// TIA Portal project "maupTIA_DEMO2023_V17" (V17)

(* hardware
DEVICE "S71500/ET200MP station_1"  S7-1500 station
   slot 0: "Rail_0"  Rack  6ES7 590-1***0-0AA0
   slot 1: "PLC_1"  CPU 1512C-1 PN  6ES7 512-1CK00-0AB0  V2.1
      slot 3: "CPU display_1"  6ES7591-1AA00-0AA0
DEVICE "HMI_1"  TP700 Comfort
   slot 0: "TP700 Comfort"  TP700 Comfort  6AV2 124-0GC01-0AX0  14.0.1.0
   slot 1: "HMI_RT_1"  TP700 Comfort  6AV2 124-0GC01-0AX0  14.0.1.0
   slot 5: "HMI_1.IE_CP_1"  PROFINET Interface  14.0.1.0
      slot 1: "PROFINET Interface_1"  PROFINET Interface
         slot 1: "Port_1"  Port
         slot 2: "Port_2"  Port
   slot 7: "HMI_1.MPI/DP_CP_1"  MPI/DP Interface  14.0.1.0
*)

// ===== PLC "PLC_1"  CPU 1512C-1 PN =====

VAR_GLOBAL   // PLC tag table "Default tag table"
   "System_Byte" AT %MB1 : Byte;
   "FirstScan" AT %M1.0 : Bool;
   "DiagStatusUpdate" AT %M1.1 : Bool;
   "AlwaysTRUE" AT %M1.2 : Bool;
   "AlwaysFALSE" AT %M1.3 : Bool;
   "Clock_Byte" AT %MB0 : Byte;
   "Clock_10Hz" AT %M0.0 : Bool;
   "Clock_5Hz" AT %M0.1 : Bool;
   "Clock_2.5Hz" AT %M0.2 : Bool;
   "Clock_2Hz" AT %M0.3 : Bool;
   "Clock_1.25Hz" AT %M0.4 : Bool;
   "Clock_1Hz" AT %M0.5 : Bool;
   "Clock_0.625Hz" AT %M0.6 : Bool;
   "Clock_0.5Hz" AT %M0.7 : Bool;
END_VAR

VAR_GLOBAL   // PLC tag table "IO"
   "diVlaveFill_Open" AT %I320.0 : Bool;
   "diVlaveFill_Close" AT %I320.1 : Bool;
   "diVlaveFill_Error" AT %I320.2 : Bool;
   "diVlaveDrain_Open" AT %I320.3 : Bool;
   "diVlaveDrain_Close" AT %I320.4 : Bool;
   "diVlaveDrain_Error" AT %I320.5 : Bool;
   "diMixer_Run" AT %I320.6 : Bool;
   "diMixer_Error" AT %I320.7 : Bool;
   "doValveFill_Open" AT %Q360.0 : Bool;
   "doValveFill_Close" AT %Q360.1 : Bool;
   "doValveDrain_Open" AT %Q360.2 : Bool;
   "doValveDrain_Close" AT %Q360.3 : Bool;
   "doMixer_Run" AT %Q360.4 : Bool;
   "aiWaterLevel" AT %IW340 : Int;
   "aoHeatPower" AT %QW380 : Int;
   "doHeatingEnable" AT %Q360.5 : Bool;
   "aiWaterTemp" AT %IW342 : Int;
END_VAR

// folder: MAUP

TYPE "Valve"
   STRUCT
      State : Struct
         Open : Bool;
         Closed : Bool;
         OpenOut : Bool;
         CloseOut : Bool;
         Err : Bool;
         StartUpFail : Bool;
         AutCtrl : Bool;
         ManCtrl : Bool;
         MayRun : Bool;
         MayAutoRun : Bool;
         GenErr : Bool;
         StColor : Int;
      END_STRUCT;
      Cmd : Struct
         AutCtrl : Bool;
         ManCtrl : Bool;
         OpenMan : Bool;
         StopMan : Bool;
         CloseMan : Bool;
         Req2OpenAut : Bool;
         Req2CloseAut : Bool;
         ResetSUF : Bool;
      END_STRUCT;
      Param : Struct
         Time2Open : Time := t#3s;
      END_STRUCT;
   END_STRUCT;
END_TYPE

TYPE "Engine"
   STRUCT
      State : Struct
         RT : DInt;
         Run : Bool;
         RunOut : Bool;
         Err : Bool;
         StartUpFail : Bool;
         AutCtrl : Bool;
         ManCtrl : Bool;
         MayRun : Bool;
         MayAutoRun : Bool;
         GenErr : Bool;
         StateInt : Int;
      END_STRUCT;
      Cmd : Struct
         SetRT : DInt := -1;
         AutCtrl : Bool;
         ManCtrl : Bool;
         TurnOnMan : Bool;
         TurnOffMan : Bool;
         Req2RunAutCtrl : Bool;
         ResetSUF : Bool;
      END_STRUCT;
      Param : Struct
         Time2Start : Time := T#3s;
      END_STRUCT;
   END_STRUCT;
END_TYPE

TYPE "Tank"
   STRUCT
      ValveFill : "Valve";
      ValveDrain : "Valve";
      Mixer : "Engine";
      Heater : "Heater";
      Draining : "PhaseDraining";
      Filling : "PhaseFilling";
      Heating : "PhaseHeating";
      Mixing : "PhaseMixing";
      GlobalError : Bool;
      WaterTemp : "AI";
      WaterLevel : "AI";
   END_STRUCT;
END_TYPE

TYPE "PhaseMixing"
   STRUCT
      Cmd : Struct
         StartAut : Bool;
         StopAut : Bool;
         StartMan : Bool;
         StopMan : Bool;
         PauseMan : Bool;
         ResumeMan : Bool;
         ResetDone : Bool;
         AutCtrl : Bool;
         ManCtrl : Bool;
      END_STRUCT;
      State : Struct
         Running : Bool;
         Idle : Bool;
         Paused : Bool;
         Done : Bool;
         AutCtrl : Bool;
         ManCtrl : Bool;
         StateInt : Int;
      END_STRUCT;
      Param : Struct
         TimeSec : Int;
      END_STRUCT;
   END_STRUCT;
END_TYPE

TYPE "PhaseFilling"
   STRUCT
      Cmd : Struct
         StartAut : Bool;
         StopAut : Bool;
         StartMan : Bool;
         StopMan : Bool;
         PauseMan : Bool;
         ResumeMan : Bool;
         ResetDone : Bool;
         AutCtrl : Bool;
         ManCtrl : Bool;
      END_STRUCT;
      State : Struct
         Running : Bool;
         Idle : Bool;
         Paused : Bool;
         Done : Bool;
         AutCtrl : Bool;
         ManCtrl : Bool;
         Stateint : Int;
      END_STRUCT;
      Param : Struct
         FillLevel : Real;
      END_STRUCT;
      WaterLevel : Real;
   END_STRUCT;
END_TYPE

TYPE "PhaseDraining"
   STRUCT
      Cmd : Struct
         StartAut : Bool;
         StopAut : Bool;
         StartMan : Bool;
         StopMan : Bool;
         PauseMan : Bool;
         ResumeMan : Bool;
         ResetDone : Bool;
         AutCtrl : Bool;
         ManCtrl : Bool;
      END_STRUCT;
      State : Struct
         Running : Bool;
         Idle : Bool;
         Paused : Bool;
         Done : Bool;
         AutCtrl : Bool;
         ManCtrl : Bool;
         StateInt : Int;
      END_STRUCT;
      Param : Struct
         DrainLevel : Real;
      END_STRUCT;
      WaterLevel : Real;
   END_STRUCT;
END_TYPE

TYPE "PhaseHeating"
   STRUCT
      Cmd : Struct
         StartAut : Bool;
         StopAut : Bool;
         StartMan : Bool;
         StopMan : Bool;
         PauseMan : Bool;
         ResumeMan : Bool;
         ResetDone : Bool;
         AutCtrl : Bool;
         ManCtrl : Bool;
      END_STRUCT;
      State : Struct
         Running : Bool;
         Idle : Bool;
         Paused : Bool;
         Done : Bool;
         AutCtrl : Bool;
         ManCtrl : Bool;
         StateInt : Int;
      END_STRUCT;
      Param : Struct
         ReqTemp : Real;
      END_STRUCT;
      WaterTemp : Real;
   END_STRUCT;
END_TYPE

TYPE "AI"
   STRUCT
      AIScaled : Real;
      TransducerLoLevel : Int;
      TransducerHiLevel : Int := 27648;
      ScaledValLoLevel : Real;
      ScaledValHiLevel : Real := 100.0;
   END_STRUCT;
END_TYPE

TYPE "Heater"
   STRUCT
      State : Struct
         EnableOut : Bool;
         HeatingOut : Real;
         AutCtrl : Bool;
         ManCtrl : Bool;
         StateInt : Int;
      END_STRUCT;
      Cmd : Struct
         AutCtrl : Bool;
         ManCtrl : Bool;
         TurnOnMan : Bool;
         TurnOffMan : Bool;
         Req2RunAutCtrl : Bool;
      END_STRUCT;
      Param : Struct
         HeatingPowerManual : Real;
         HeatingSetPointAutomat : Real;
      END_STRUCT;
   END_STRUCT;
END_TYPE

// folder: (top level)

DATA_BLOCK "TankFC_DB"   // DB4
{ S7_Optimized_Access := 'TRUE' }
VERSION : 0.1
// stored: InstanceOfName TankFC
"TankFC"
BEGIN
END_DATA_BLOCK

// folder: DBs

DATA_BLOCK "Data"   // DB1
{ S7_Optimized_Access := 'TRUE' }
VERSION : 0.1
   VAR
      Tank1 : "Tank";
   END_VAR
BEGIN
   Tank1.Filling.Param.FillLevel := 1.95;
   Tank1.ValveDrain.Param.Time2Open := T#30m;
   Tank1.ValveFill.Param.Time2Open := T#30m;
   Tank1.Mixer.Param.Time2Start := T#30m;
   Tank1.WaterTemp.ScaledValLoLevel := 0.0;
   Tank1.WaterTemp.ScaledValHiLevel := 100.0;
   Tank1.WaterLevel.ScaledValHiLevel := 2.0;
   Tank1.Mixing.Param.TimeSec := 10;
   Tank1.Heating.Param.ReqTemp := 95.0;
   Tank1.Heater.Param.HeatingPowerManual := 0.0;
END_DATA_BLOCK

// folder: System blocks/Program resources

DATA_BLOCK "IsTime2Open"   // DB2
{ S7_Optimized_Access := 'TRUE' }
AUTHOR : Simatic
FAMILY : IEC
NAME : IEC_TMR
VERSION : 1.0
// stored: InstanceOfName IEC_TIMER
"IEC_TIMER"
BEGIN
END_DATA_BLOCK

DATA_BLOCK "IsReallyRunning"   // DB6
{ S7_Optimized_Access := 'TRUE' }
AUTHOR : Simatic
FAMILY : IEC
NAME : IEC_TMR
VERSION : 1.0
// stored: InstanceOfName IEC_TIMER
"IEC_TIMER"
BEGIN
END_DATA_BLOCK

DATA_BLOCK "IsTime2Close"   // DB7
{ S7_Optimized_Access := 'TRUE' }
AUTHOR : Simatic
FAMILY : IEC
NAME : IEC_TMR
VERSION : 1.0
// stored: InstanceOfName IEC_TIMER
"IEC_TIMER"
BEGIN
END_DATA_BLOCK

// folder: (top level)

FUNCTION_BLOCK "TankFC"   // FB3, LAD
{ S7_Optimized_Access := 'TRUE' }
VERSION : 0.1
   VAR_INPUT
      diMixer_Running : Bool;
      diMixer_Error : Bool;
      diValveFill_Open : Bool;
      diValveFill_Close : Bool;
      diValveFill_Error : Bool;
      diValveDrain_Open : Bool;
      diValveDrain_Close : Bool;
      diValveDrain_Error : Bool;
      aiWaterLevel : Int;
      aiWaterTemp : Int;
   END_VAR
   VAR_OUTPUT
      doMixerStart : Bool;
      doValveFill_Open : Bool;
      doValveFill_Close : Bool;
      doValveDrain_Open : Bool;
      doValveDrain_Close : Bool;
      doHeatingEnable : Bool;
      aoReqPowerOfHeating : Word;
   END_VAR
   VAR_IN_OUT
      Tank : "Tank";
   END_VAR
   VAR
      Mixer : "Eng_1DO";
      ValveFill : "Val_2DO";
      ValveDrain : "Val_2DO";
      DrainingFC_Instance : "DrainingFC";
      FillingFC_Instance : "FillingFC";
      MixingFC_Instance : "MixingFC";
      Real2AnalogValue_Instance : "Real2AnalogValue";
      HeatingFC_Instance : "HeatingFC";
      HeaterFC_Instance : "HeaterFC";
   END_VAR
   VAR_TEMP
      HeaterReqPower : Real;
   END_VAR
   VAR_TEMP   // added for the SCL form of the ladder/FBD networks
      _w1 : Bool;
      _w2 : Bool;
   END_VAR
BEGIN

REGION Network 1
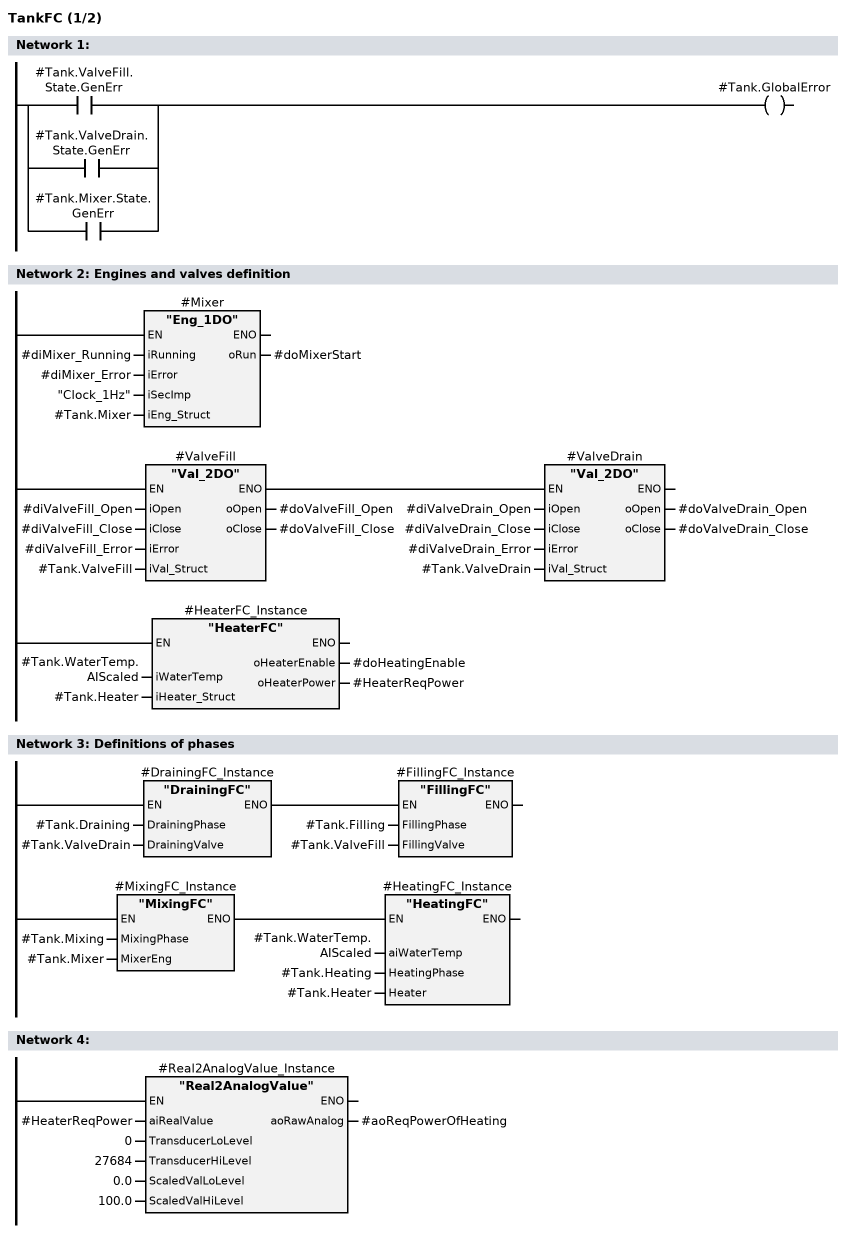
   RUNG wire#powerrail
      Contact( #Tank.ValveFill.State.GenErr )
      wire#w1
      Coil( #Tank.GlobalError )
   END_RUNG
   RUNG wire#powerrail
      Contact( #Tank.ValveDrain.State.GenErr )
   END_RUNG wire#w1
   RUNG wire#powerrail
      Contact( #Tank.Mixer.State.GenErr )
   END_RUNG wire#w1
   // the same network as SCL:
   #Tank.GlobalError := #Tank.ValveFill.State.GenErr OR #Tank.ValveDrain.State.GenErr OR #Tank.Mixer.State.GenErr;
END_REGION

REGION Network 2: Engines and valves definition
   RUNG wire#powerrail
      #Mixer(iRunning := #diMixer_Running, iError := #diMixer_Error, iSecImp := "Clock_1Hz", iEng_Struct := #Tank.Mixer, oRun => #doMixerStart)
   END_RUNG
   RUNG wire#powerrail
      #ValveFill(iOpen := #diValveFill_Open, iClose := #diValveFill_Close, iError := #diValveFill_Error, iVal_Struct := #Tank.ValveFill, oOpen => #doValveFill_Open, oClose => #doValveFill_Close)
      #ValveDrain(iOpen := #diValveDrain_Open, iClose := #diValveDrain_Close, iError := #diValveDrain_Error, iVal_Struct := #Tank.ValveDrain, oOpen => #doValveDrain_Open, oClose => #doValveDrain_Close)
   END_RUNG
   RUNG wire#powerrail
      #HeaterFC_Instance(iWaterTemp := #Tank.WaterTemp.AIScaled, iHeater_Struct := #Tank.Heater, oHeaterEnable => #doHeatingEnable, oHeaterPower => #HeaterReqPower)
   END_RUNG
   // the same network as SCL:
   #Mixer(iRunning := #diMixer_Running,   // "Eng_1DO"
          iError := #diMixer_Error,
          iSecImp := "Clock_1Hz",
          iEng_Struct := #Tank.Mixer,
          oRun => #doMixerStart);
   #ValveFill(iOpen := #diValveFill_Open,   // "Val_2DO"
              iClose := #diValveFill_Close,
              iError := #diValveFill_Error,
              iVal_Struct := #Tank.ValveFill,
              oOpen => #doValveFill_Open,
              oClose => #doValveFill_Close,
              ENO => #_w1);
   IF #_w1 THEN
       #ValveDrain(iOpen := #diValveDrain_Open,   // "Val_2DO"
                   iClose := #diValveDrain_Close,
                   iError := #diValveDrain_Error,
                   iVal_Struct := #Tank.ValveDrain,
                   oOpen => #doValveDrain_Open,
                   oClose => #doValveDrain_Close);
   END_IF;
   #HeaterFC_Instance(iWaterTemp := #Tank.WaterTemp.AIScaled,   // "HeaterFC"
                      iHeater_Struct := #Tank.Heater,
                      oHeaterEnable => #doHeatingEnable,
                      oHeaterPower => #HeaterReqPower);
END_REGION

REGION Network 3: Definitions of phases
   RUNG wire#powerrail
      #DrainingFC_Instance(DrainingPhase := #Tank.Draining, DrainingValve := #Tank.ValveDrain)
      #FillingFC_Instance(FillingPhase := #Tank.Filling, FillingValve := #Tank.ValveFill)
   END_RUNG
   RUNG wire#powerrail
      #MixingFC_Instance(MixingPhase := #Tank.Mixing, MixerEng := #Tank.Mixer)
      #HeatingFC_Instance(aiWaterTemp := #Tank.WaterTemp.AIScaled, HeatingPhase := #Tank.Heating, Heater := #Tank.Heater)
   END_RUNG
   // the same network as SCL:
   #DrainingFC_Instance(DrainingPhase := #Tank.Draining, DrainingValve := #Tank.ValveDrain, ENO => #_w1);   // "DrainingFC"
   IF #_w1 THEN
       #FillingFC_Instance(FillingPhase := #Tank.Filling, FillingValve := #Tank.ValveFill);   // "FillingFC"
   END_IF;
   #MixingFC_Instance(MixingPhase := #Tank.Mixing, MixerEng := #Tank.Mixer, ENO => #_w2);   // "MixingFC"
   IF #_w2 THEN
       #HeatingFC_Instance(aiWaterTemp := #Tank.WaterTemp.AIScaled,   // "HeatingFC"
                           HeatingPhase := #Tank.Heating,
                           Heater := #Tank.Heater);
   END_IF;
END_REGION

REGION Network 4
   RUNG wire#powerrail
      #Real2AnalogValue_Instance(aiRealValue := #HeaterReqPower, TransducerLoLevel := 0, TransducerHiLevel := 27684, ScaledValLoLevel := 0.0, ScaledValHiLevel := 100.0, aoRawAnalog => #aoReqPowerOfHeating)
   END_RUNG
   // the same network as SCL:
   #Real2AnalogValue_Instance(aiRealValue := #HeaterReqPower,   // "Real2AnalogValue"
                           TransducerLoLevel := 0,
                           TransducerHiLevel := 27684,
                           ScaledValLoLevel := 0.0,
                           ScaledValHiLevel := 100.0,
                           aoRawAnalog => #aoReqPowerOfHeating);
END_REGION

REGION Network 5: Analog scaling
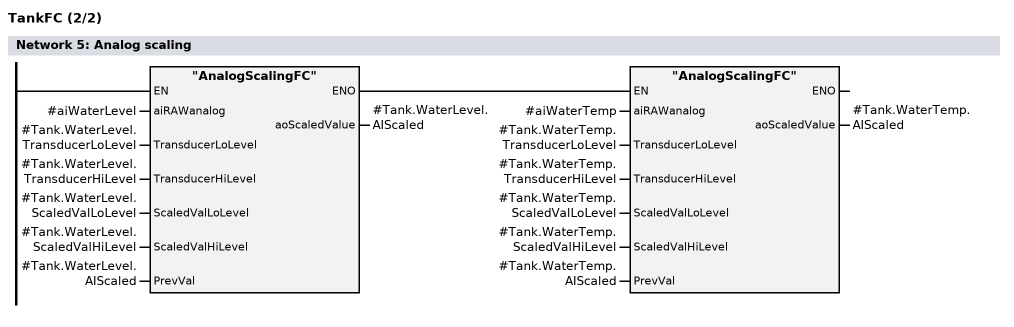
   RUNG wire#powerrail
      "AnalogScalingFC"(aiRAWanalog := #aiWaterLevel, TransducerLoLevel := #Tank.WaterLevel.TransducerLoLevel, TransducerHiLevel := #Tank.WaterLevel.TransducerHiLevel, ScaledValLoLevel := #Tank.WaterLevel.ScaledValLoLevel, ScaledValHiLevel := #Tank.WaterLevel.ScaledValHiLevel, PrevVal := #Tank.WaterLevel.AIScaled, aoScaledValue => #Tank.WaterLevel.AIScaled)
      "AnalogScalingFC"(aiRAWanalog := #aiWaterTemp, TransducerLoLevel := #Tank.WaterTemp.TransducerLoLevel, TransducerHiLevel := #Tank.WaterTemp.TransducerHiLevel, ScaledValLoLevel := #Tank.WaterTemp.ScaledValLoLevel, ScaledValHiLevel := #Tank.WaterTemp.ScaledValHiLevel, PrevVal := #Tank.WaterTemp.AIScaled, aoScaledValue => #Tank.WaterTemp.AIScaled)
   END_RUNG
   // the same network as SCL:
   "AnalogScalingFC"(aiRAWanalog := #aiWaterLevel,
                     TransducerLoLevel := #Tank.WaterLevel.TransducerLoLevel,
                     TransducerHiLevel := #Tank.WaterLevel.TransducerHiLevel,
                     ScaledValLoLevel := #Tank.WaterLevel.ScaledValLoLevel,
                     ScaledValHiLevel := #Tank.WaterLevel.ScaledValHiLevel,
                     PrevVal := #Tank.WaterLevel.AIScaled,
                     aoScaledValue => #Tank.WaterLevel.AIScaled,
                     ENO => #_w1);
   IF #_w1 THEN
       "AnalogScalingFC"(aiRAWanalog := #aiWaterTemp,
                         TransducerLoLevel := #Tank.WaterTemp.TransducerLoLevel,
                         TransducerHiLevel := #Tank.WaterTemp.TransducerHiLevel,
                         ScaledValLoLevel := #Tank.WaterTemp.ScaledValLoLevel,
                         ScaledValHiLevel := #Tank.WaterTemp.ScaledValHiLevel,
                         PrevVal := #Tank.WaterTemp.AIScaled,
                         aoScaledValue => #Tank.WaterTemp.AIScaled);
   END_IF;
END_REGION

REGION Network 6 (SCL): Data transfer
   #Tank.Draining.WaterLevel := #Tank.WaterLevel.AIScaled;
   #Tank.Filling.WaterLevel := #Tank.WaterLevel.AIScaled;
   #Tank.Heating.WaterTemp := #Tank.WaterTemp.AIScaled;
END_REGION
END_FUNCTION_BLOCK

ORGANIZATION_BLOCK "Main"   // OB1, LAD, ProgramCycle
TITLE = "Main Program Sweep (Cycle)"
{ S7_Optimized_Access := 'TRUE' }
VERSION : 0.1
   VAR_INPUT
      Initial_Call : Bool;   // Initial call of this OB
      Remanence : Bool;   // =True, if remanent data are available
   END_VAR
BEGIN
END_ORGANIZATION_BLOCK

ORGANIZATION_BLOCK "Cyclic interrupt10ms"   // OB31, LAD, CyclicInterrupt
{ S7_Optimized_Access := 'TRUE' }
VERSION : 0.1
   VAR_INPUT
      Initial_Call : Bool;   // Initial call of this OB
      Event_Count : Int;   // Events discarded
   END_VAR
BEGIN

REGION Network 1
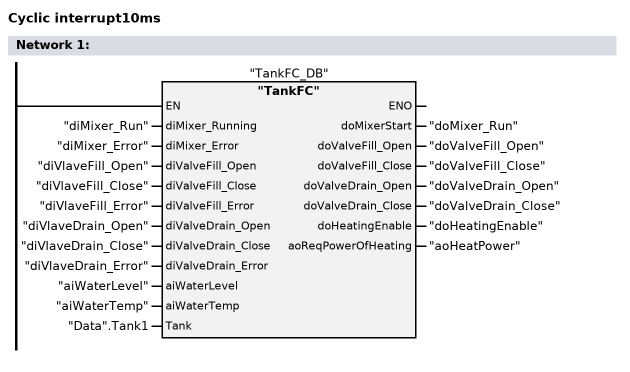
   RUNG wire#powerrail
      "TankFC_DB"(diMixer_Running := "diMixer_Run", diMixer_Error := "diMixer_Error", diValveFill_Open := "diVlaveFill_Open", diValveFill_Close := "diVlaveFill_Close", diValveFill_Error := "diVlaveFill_Error", diValveDrain_Open := "diVlaveDrain_Open", diValveDrain_Close := "diVlaveDrain_Close", diValveDrain_Error := "diVlaveDrain_Error", aiWaterLevel := "aiWaterLevel", aiWaterTemp := "aiWaterTemp", Tank := "Data".Tank1, doMixerStart => "doMixer_Run", doValveFill_Open => "doValveFill_Open", doValveFill_Close => "doValveFill_Close", doValveDrain_Open => "doValveDrain_Open", doValveDrain_Close => "doValveDrain_Close", doHeatingEnable => "doHeatingEnable", aoReqPowerOfHeating => "aoHeatPower")
   END_RUNG
   // the same network as SCL:
   "TankFC_DB"(diMixer_Running := "diMixer_Run",   // "TankFC"
               diMixer_Error := "diMixer_Error",
               diValveFill_Open := "diVlaveFill_Open",
               diValveFill_Close := "diVlaveFill_Close",
               diValveFill_Error := "diVlaveFill_Error",
               diValveDrain_Open := "diVlaveDrain_Open",
               diValveDrain_Close := "diVlaveDrain_Close",
               diValveDrain_Error := "diVlaveDrain_Error",
               aiWaterLevel := "aiWaterLevel",
               aiWaterTemp := "aiWaterTemp",
               Tank := "Data".Tank1,
               doMixerStart => "doMixer_Run",
               doValveFill_Open => "doValveFill_Open",
               doValveFill_Close => "doValveFill_Close",
               doValveDrain_Open => "doValveDrain_Open",
               doValveDrain_Close => "doValveDrain_Close",
               doHeatingEnable => "doHeatingEnable",
               aoReqPowerOfHeating => "aoHeatPower");
END_REGION
END_ORGANIZATION_BLOCK

ORGANIZATION_BLOCK "Startup"   // OB100, SCL, Startup
TITLE = "Complete Restart"
{ S7_Optimized_Access := 'TRUE' }
VERSION : 0.1
   VAR_INPUT
      LostRetentive : Bool;   // True if retentive data are lost
      LostRTC : Bool;   // True if date and time are lost
   END_VAR
BEGIN
END_ORGANIZATION_BLOCK

// folder: FCs

FUNCTION_BLOCK "Eng_1DO"   // FB1, SCL
{ S7_Optimized_Access := 'TRUE' }
VERSION : 0.1
   VAR_INPUT
      iRunning : Bool;
      iError : Bool;
      iSecImp : Bool;
   END_VAR
   VAR_OUTPUT
      oRun : Bool;
   END_VAR
   VAR_IN_OUT
      iEng_Struct : "Engine";
   END_VAR
   VAR
      SecImpEdge : R_TRIG;
      SUF_Timer : TON_TIME;
   END_VAR
   VAR_TEMP
      Rising_Edge : Bool;
      TimerDone : Bool;
   END_VAR
   VAR CONSTANT
      Running : Int := 0;
      Stop : Int := 1;
      RunningAndErr : Int := 2;
      Err : Int := 3;
   END_VAR
BEGIN
   REGION RunningTime  
       // counting running time of engine - (motoseconds in real situation it should be moto hours)
       // detection rising edge of input secimp - should be conected 1Hz internal clock from PLC

       // je zpetna vazba od zarizeni kladna?
       IF #iEng_Struct.State.Run THEN
           // detekce nabezne hrany pomoci bit. logic. oper. R_TRIG
           "SecImpEdge"(CLK := "Clock_1Hz",
                        Q => #Rising_Edge); // pridani Rising_Edge {bool} do Temp

           // detekce nabezne hrany
           IF #Rising_Edge = TRUE THEN
               #iEng_Struct.State.RT := #iEng_Struct.State.RT + 1; // inkrementace motohodin
               #Rising_Edge := FALSE; // resetovani nabezne hrany
               ;
           END_IF;

           // uzivatelske nastaveni motosekund
           IF #iEng_Struct.Cmd.SetRT >= 0 THEN
               #iEng_Struct.State.RT := #iEng_Struct.Cmd.SetRT; // zmena  motohodin na zadanou hodnotu commandem;
               #iEng_Struct.Cmd.SetRT := -1; // zmena setRT na -1
           END_IF;
           ;
       END_IF;

   END_REGION

   REGION RunState 
       // set real state of engine input into engine structure - input of running
       // engine can be taken from frequential converter, speed sensor, or just
       // from switching element
       // 
       // Zda zařízení skutečně běží, není možné určit pouze tím, že jsme zadali příkaz k
       //jeho sepnutí. DO stavu Run tedy nastavte hodnotu vyčtenou ze zpětné vazby od
       //zařízení (#iRunning).

       #iEng_Struct.State.Run := #iRunning;

   END_REGION

   REGION Manual/Automat 
       // switching state of engine - automatic or manual control (default state is manual)

       IF #iEng_Struct.Cmd.AutCtrl THEN
           // Automaticky rezim
           #iEng_Struct.State.AutCtrl := TRUE;
           #iEng_Struct.State.ManCtrl := FALSE;
           #iEng_Struct.Cmd.ManCtrl := FALSE;
           #iEng_Struct.Cmd.AutCtrl := FALSE;
       END_IF;

       IF #iEng_Struct.Cmd.ManCtrl THEN
           // Manualni rezim (preferovaný, pokud není aktivní automatický režim)
           #iEng_Struct.State.AutCtrl := FALSE;
           #iEng_Struct.State.ManCtrl := TRUE;
           #iEng_Struct.Cmd.ManCtrl := FALSE;
           #iEng_Struct.Cmd.AutCtrl := FALSE;
       END_IF;

       IF #iEng_Struct.State.ManCtrl = FALSE AND #iEng_Struct.State.AutCtrl = FALSE THEN
           // preferovaný MANUALNI, pokud není aktivní automatický režim)
           #iEng_Struct.State.AutCtrl := FALSE;
           #iEng_Struct.State.ManCtrl := TRUE;
       END_IF;

       // Resetovani prikazu po provedeni zmen
       #iEng_Struct.Cmd.AutCtrl := FALSE;
       #iEng_Struct.Cmd.ManCtrl := FALSE;

   END_REGION

   REGION MR/MAR 
       // setting auxilary signals (may run, may auto run) - MR AND NOT MAR - eng should be started in manual mode,
       // MAR - should be started in automatic mode

       IF #iEng_Struct.State.ManCtrl AND #iEng_Struct.State.Err = FALSE THEN
           // MayRun je aktivni
           #iEng_Struct.State.MayRun := TRUE;
           #iEng_Struct.State.MayAutoRun := FALSE;
       END_IF;

       IF #iEng_Struct.State.AutCtrl AND #iEng_Struct.State.Err = FALSE THEN
           // MayAutoRun je aktivni
           #iEng_Struct.State.MayAutoRun := TRUE;
           #iEng_Struct.State.MayRun := FALSE;
       END_IF;

   END_REGION

   REGION ManCtrl
       // processing manual actions - if command is processed, it is set to FALSE even if can't be processed
       // Engine commands are turn off (stop) and turn on (start)

       IF #iEng_Struct.Cmd.TurnOnMan AND #iEng_Struct.State.MayRun THEN
           // aktivace stavu RunOut
           #iEng_Struct.State.RunOut := TRUE;
           #iEng_Struct.Cmd.TurnOnMan := FALSE;
       END_IF;

       IF #iEng_Struct.Cmd.TurnOffMan AND #iEng_Struct.State.MayRun THEN
           // deaktivace stavu RunOut
           #iEng_Struct.State.RunOut := FALSE;
           #iEng_Struct.Cmd.TurnOffMan := FALSE;
       END_IF;


       // vynulovani obou prikazu


   END_REGION

   REGION AutCtrl 
       //if request to run in automatic mode set outputs to right states if MAR
       //AutoRequest shouldn't be reseted to false state

       IF #iEng_Struct.State.AutCtrl AND #iEng_Struct.State.MayAutoRun THEN
           // otestujte příkaz Req2RunAutCtrl. Na základě jeho hodnoty nastavte opět stav RunOut.
           #iEng_Struct.State.RunOut := #iEng_Struct.Cmd.Req2RunAutCtrl;
       END_IF;

   END_REGION


   REGION ErrStates
       // definition of error states 
       // error - input from digital input of plc - fyzical state of engine 
       // calculating start up fail - if output is sets to start engine, it's expected feedback from running signal in defined time, if feedback doesn't show in this time, it should be start up fail error
       // merge of these two error is general error

       // timer se aktivuje pokud je odeslan prikaz na spusteni motoru, pokud do doby Time2Start neprijde iRunning = TRUE, tak se TimerDone = TRUE 
       // Pridan TimerDone do Temp{}
       "IsReallyRunning".TON(IN := #iEng_Struct.State.Run,
                             PT := #iEng_Struct.Param.Time2Start,
                             Q => #TimerDone);

       IF #TimerDone AND #iRunning = FALSE THEN
           // Pokud do této doby není aktivní zpětná vazba od zařízení, vygeneruje se příznak (stav) StartUpFail.
           #iEng_Struct.State.StartUpFail := TRUE;
       END_IF;

       IF #TimerDone = FALSE AND #iRunning THEN
           // Resetovani chyby -> timer neni done ale prisla zpetna vazba, ze motor bezi
           #iEng_Struct.State.StartUpFail := FALSE;
       END_IF;

       IF #iError THEN
           // pokud zařízení aktivovalo svůj výstup iError (vstup do PLC), nastavte příznak (stav) #Err
           #iEng_Struct.State.Err := TRUE;
       ELSE
           #iEng_Struct.State.Err := FALSE;
       END_IF;

       //Logickým součtem obou výše popsaných chybových příznaků je příznak GenErr.
       #iEng_Struct.State.GenErr := #iEng_Struct.State.StartUpFail OR #iEng_Struct.State.Err;

       IF #iEng_Struct.Cmd.ResetSUF THEN
           // Příkaz ResetSUF resetuje příznak StartUpFail. Nezapomeňte vyresetovat i tento příkaz!
           #iEng_Struct.State.GenErr := FALSE;
           #iEng_Struct.Cmd.ResetSUF := FALSE;
       END_IF;

       IF #iEng_Struct.State.GenErr THEN
           // Pokud je aktivní příznak GenErr, je nutné vypnout výstup modulu (deaktivovat zařízení - přepnout DO bezpečného stavu) - RunOut.
           #iEng_Struct.State.RunOut := TRUE;
       END_IF;




   END_REGION
   (*
   Za blok ErrStates vložte příkaz, který zrcadlí hodnotu stavu RunOut z
   datového bloku na výstup #oRun. Hodnoty jsou duplikovány, protože
   zatímco RunOut je možné i číst a je využívána ve vizualizaci, výstup oRun
   je připojen přes výstup funkčního bloku tanku přímo na fyzický výstup
   PLC a ovládá zařízení.
   *)
   #oRun := #iEng_Struct.State.RunOut;

   REGION StatusInt
       //write combination of states into int value for visualization (engine - combination of running state and error)
       //

       IF #iEng_Struct.State.GenErr = FALSE AND #iEng_Struct.State.Run THEN
           // Pokud není GenErr a modul je spuštěn (ve stavu Run), přiřaďte konstantu #Running (0)
           #iEng_Struct.State.StateInt := #Running;
       END_IF;

       IF #iEng_Struct.State.GenErr = FALSE AND #iEng_Struct.State.Run = FALSE THEN //NEJSEM SI JIST PODMINKOIU, KDZY MODUL JE ZASTAVEN
           // Pokud není GenErr a modul je zastaven, přiřaďte konstantu #Stop (1)
           #iEng_Struct.State.StateInt := #Stop;
       END_IF;

       IF #iEng_Struct.State.GenErr THEN
           // Pokud je GenErr, nastavte na základě stavu Run konstanty #RunningAndErr (2) nebo pouze #Err (3).
           IF #iEng_Struct.State.Run THEN
               #iEng_Struct.State.StateInt := #RunningAndErr;
           ELSE
               #iEng_Struct.State.StateInt := #Err;
           END_IF;
           ;
       END_IF;


   END_REGION
END_FUNCTION_BLOCK

FUNCTION_BLOCK "Val_2DO"   // FB2, SCL
{ S7_Optimized_Access := 'TRUE' }
VERSION : 0.1
   VAR_INPUT
      iOpen : Bool;
      iClose : Bool;
      iError : Bool;
   END_VAR
   VAR_OUTPUT
      oOpen : Bool;
      oClose : Bool;
   END_VAR
   VAR_IN_OUT
      iVal_Struct : "Valve";
   END_VAR
   VAR
      fTimeToOpen : TON_TIME;
      fTimeToClose : TON_TIME;
   END_VAR
   VAR_TEMP
      Ton_1_starter : Bool;
      Ton_1_done : Bool;
      Ton_2_starter : Bool;
      Ton_2_done : Bool;
   END_VAR
   VAR CONSTANT
      Open : Int := 0;
      Closed : Int := 1;
      OpenAndErr : Int := 2;
      ClosedAndErr : Int := 3;
      NotOpenNotClosedNotErr : Int := 4;
      NotOpenNotClosedAndErr : Int := 5;
      OpenAndClosedAndErr : Int := 6;
      OpenAndClosedNotErr : Int := 7;
   END_VAR
BEGIN
   REGION OpenState 
       // set real state of valve input into valve structure - input of valve can be taken from limit sensor...

       // NEJSEM SI TIMTO JIST
       #iVal_Struct.State.Open := #iOpen;
       #iVal_Struct.State.Closed := #iClose;

   END_REGION

   REGION Manual/Automat
       // switching state of engine - automatic or manual control (default state is manual)

       IF #iVal_Struct.Cmd.AutCtrl THEN
           // automaticky rezim
           #iVal_Struct.State.AutCtrl := TRUE;
           #iVal_Struct.State.ManCtrl := FALSE;
           #iVal_Struct.Cmd.ManCtrl := FALSE;
       END_IF;

       IF #iVal_Struct.Cmd.ManCtrl THEN
           // manualni rezim
           #iVal_Struct.State.AutCtrl := FALSE;
           #iVal_Struct.State.ManCtrl := TRUE;
           #iVal_Struct.Cmd.AutCtrl := FALSE;
       END_IF;

       IF #iVal_Struct.State.AutCtrl = FALSE AND #iVal_Struct.State.ManCtrl = FALSE THEN
           // defaultne manual
           #iVal_Struct.State.ManCtrl := TRUE;
           #iVal_Struct.State.AutCtrl := FALSE;
       END_IF;


       // resetovani prikazu po provedeni zmen
       #iVal_Struct.Cmd.AutCtrl := FALSE;
       #iVal_Struct.Cmd.ManCtrl := FALSE;

   END_REGION

   REGION MR/MAR
       // setting auxilary signals (may run, may auto run) - MR AND NOT MAR - eng should be started in manual mode, MAR - should be started in automatic mode
       IF #iVal_Struct.State.ManCtrl AND #iVal_Struct.State.Err = FALSE THEN
           // MayRun je aktivni
           #iVal_Struct.State.MayRun := TRUE;
           #iVal_Struct.State.MayAutoRun := FALSE;
       END_IF;

       IF #iVal_Struct.State.AutCtrl AND #iVal_Struct.State.Err = FALSE THEN
           // MayAutoRun je aktivni
           #iVal_Struct.State.MayAutoRun := TRUE;
           #iVal_Struct.State.MayRun := FALSE;
       END_IF;

   END_REGION

   REGION ManCtrl
       // processing manual actions - if command is processed, it is sets to FALSE even if can't be processed
       // Valve commands are open, close and stop - valve can be stopped intermediate position

       IF #iVal_Struct.Cmd.OpenMan AND #iVal_Struct.State.MayRun THEN
           // Pokud je aktivní příkaz OpenMan a současně je aktivní pomocný příznak pro
           // manuální režim, aktivujte stav OpenOut a deaktivujte stav CloseOut.
           #iVal_Struct.State.OpenOut := TRUE;
           #iVal_Struct.State.CloseOut := FALSE;
       END_IF;

       IF #iVal_Struct.Cmd.CloseMan AND #iVal_Struct.State.MayRun THEN
           // Deaktivace openout a aktivace closeout
           #iVal_Struct.State.OpenOut := FALSE;
           #iVal_Struct.State.CloseOut := TRUE;
       END_IF;

       IF #iVal_Struct.Cmd.StopMan THEN
           // deaktivace obou stavu
           #iVal_Struct.State.OpenOut := FALSE;
           #iVal_Struct.State.CloseOut := FALSE;
       END_IF;

       // VYNULOVANI PRIKAZU
       #iVal_Struct.Cmd.OpenMan := FALSE;
       #iVal_Struct.Cmd.StopMan := FALSE;
       #iVal_Struct.Cmd.CloseMan := FALSE;

   END_REGION

   REGION AutCtrl
       //if request to run in automatic mode -> set outputs to right states if MAR
       //AutoRequest shouldn't be reseted to false state
       //if request to open and request to close are setted to 1 simultaneously - outputs should be 0.

       IF #iVal_Struct.State.AutCtrl AND #iVal_Struct.State.MayAutoRun THEN
           // Statement section IF
           IF #iVal_Struct.Cmd.Req2OpenAut AND #iVal_Struct.Cmd.Req2CloseAut = FALSE THEN
               // Statement section IF
               #iVal_Struct.State.OpenOut := TRUE;
               #iVal_Struct.State.CloseOut := FALSE;
           END_IF;

           IF #iVal_Struct.Cmd.Req2OpenAut = FALSE AND #iVal_Struct.Cmd.Req2CloseAut THEN
               // Statement section IF
               #iVal_Struct.State.OpenOut := FALSE;
               #iVal_Struct.State.CloseOut := TRUE;
           END_IF;

           IF #iVal_Struct.Cmd.Req2OpenAut = FALSE AND #iVal_Struct.Cmd.Req2CloseAut = FALSE THEN
               // Statement section IF
               #iVal_Struct.State.OpenOut := FALSE;
               #iVal_Struct.State.CloseOut := FALSE;
           END_IF;
       END_IF;

       // #iVal_Struct.Cmd.Req2OpenAut := FALSE;
       //#iVal_Struct.Cmd.Req2CloseAut := FALSE;

   END_REGION

   REGION ErrStates´
       // definition of error states 
       // error - input from digital input of plc - fyzical state of valve
       // calculating start up fail - if output is sets to open or close, it's expected feedback from limit sensor in defined time, if feedback doesn't show in this time, it should be start up fail error
       // merge of these two error is general error
       // error is both inputs (open and closed) true state


       // start up fail can be reseted by operator, command resetSUF, resets SUF and engine should be started again


       // if error state exists outputs should be in stop state

   (*  *)

       "IsTime2Open".TON(IN := #Ton_1_starter,
                         PT := #iVal_Struct.Param.Time2Open,
                         Q => #Ton_1_done);

       "IsTime2Close".TON(IN := #Ton_2_starter,
                          PT := #iVal_Struct.Param.Time2Open,
                          Q => #Ton_2_done);
       IF #iVal_Struct.State.OpenOut AND #iVal_Struct.State.CloseOut = FALSE THEN
           // Statement section IF
           #Ton_1_starter := TRUE;
       ELSE
           #Ton_1_starter := FALSE;
       END_IF;


       IF #Ton_1_done = FALSE THEN
           IF #iOpen = FALSE THEN
               #iVal_Struct.State.StartUpFail := #Ton_1_done OR #Ton_2_done;
           END_IF;
       END_IF;

       IF #iVal_Struct.State.OpenOut = FALSE AND #iVal_Struct.State.CloseOut THEN
           // podminka pro sepnuti casovace 1
           #Ton_2_starter := TRUE;
       ELSE
           #Ton_2_starter := FALSE;
       END_IF;

       // Pokud do doby casovace ton2 neprijde zpetna vazba od ventilu vygeneruj chybu startupfail
       // Hodnota je log soucet cystupu casovacu
       IF #Ton_2_done = FALSE THEN
           IF #iClose = FALSE THEN
               #iVal_Struct.State.StartUpFail := #Ton_1_done OR #Ton_2_done;
           END_IF;
       END_IF;

       IF #iError THEN
           #iVal_Struct.State.Err := TRUE;
       ELSE
           #iVal_Struct.State.Err := FALSE;
       END_IF;

       // GENERAL ERROR - log soucet iError & Startupfail
       #iVal_Struct.State.GenErr := #iVal_Struct.State.StartUpFail OR #iVal_Struct.State.Err;

       // reset priznaku startupfails
       IF #iVal_Struct.Cmd.ResetSUF THEN
           // Příkaz ResetSUF resetuje příznak StartUpFail. Nezapomeňte vyresetovat i tento příkaz!
           #iVal_Struct.State.GenErr := FALSE;
           #iVal_Struct.Cmd.ResetSUF := FALSE;
       END_IF;

       IF #iVal_Struct.State.GenErr THEN
           // Pokud je aktivní příznak GenErr, je nutné vypnout výstupy modulu -> prepnout do bezpecneho stavu{openout closeout}
           #iVal_Struct.State.OpenOut := TRUE;
           #iVal_Struct.State.CloseOut := TRUE;
       END_IF;


   END_REGION
   (*
   Za blok ErrStates vložte příkaz, který zrcadlí hodnotu stavů OpenOut a
   CloseOut z datového bloku na výstup #oOpen a #oClose. Hodnoty jsou
   duplikovány, protože zatímco OpenOut a CloseOut je možné i číst a je
   využívána ve vizualizaci, výstupy #oOpen a #oClose jsou připojeny přes
   výstup funkčního bloku tanku přímo na fyzické výstupy PLC a ovládají
   zařízení.
   *)
   #oOpen := #iVal_Struct.State.OpenOut;
   #oClose := #iVal_Struct.State.CloseOut;

   REGION StatusInt
       //write combination of states into int value for visualization (valve - combination of open, close state and error)
       IF #iVal_Struct.State.Open AND NOT #iVal_Struct.State.Closed AND NOT #iVal_Struct.State.GenErr THEN
           #iVal_Struct.State.StColor := #Open;
       ELSIF NOT #iVal_Struct.State.Open AND #iVal_Struct.State.Closed AND NOT #iVal_Struct.State.GenErr THEN
           #iVal_Struct.State.StColor := #Closed;
       ELSIF #iVal_Struct.State.Open AND NOT #iVal_Struct.State.Closed AND #iVal_Struct.State.GenErr THEN
           #iVal_Struct.State.StColor := #OpenAndErr;
       ELSIF NOT #iVal_Struct.State.Open AND #iVal_Struct.State.Closed AND #iVal_Struct.State.GenErr THEN
           #iVal_Struct.State.StColor := #ClosedAndErr;
       ELSIF NOT #iVal_Struct.State.Open AND NOT #iVal_Struct.State.Closed AND NOT #iVal_Struct.State.GenErr THEN
           #iVal_Struct.State.StColor := #NotOpenNotClosedNotErr;
       ELSIF NOT #iVal_Struct.State.Open AND NOT #iVal_Struct.State.Closed AND #iVal_Struct.State.GenErr THEN
           #iVal_Struct.State.StColor := #NotOpenNotClosedAndErr;
       ELSIF #iVal_Struct.State.Open AND #iVal_Struct.State.Closed AND #iVal_Struct.State.GenErr THEN
           #iVal_Struct.State.StColor := #OpenAndClosedAndErr;
       ELSIF #iVal_Struct.State.Open AND #iVal_Struct.State.Closed AND NOT #iVal_Struct.State.GenErr THEN
           #iVal_Struct.State.StColor := #OpenAndClosedNotErr;
       END_IF;
   END_REGION
END_FUNCTION_BLOCK

FUNCTION_BLOCK "FillingFC"   // FB4, SCL
{ S7_Optimized_Access := 'TRUE' }
VERSION : 0.1
   VAR_IN_OUT
      FillingPhase : "PhaseFilling";
      FillingValve : "Valve";
   END_VAR
   VAR CONSTANT
      Idle : Int := 0;
      Running : Int := 1;
      Pause : Int := 2;
   END_VAR
BEGIN
   REGION Aut/Man
       // switching state of engine - automatic or manual control (default state is manual)
       IF #FillingPhase.Cmd.AutCtrl THEN
           #FillingPhase.State.ManCtrl := FALSE;
           #FillingPhase.State.AutCtrl := TRUE;
           #FillingPhase.Cmd.AutCtrl := FALSE;
       END_IF;

       IF #FillingPhase.Cmd.ManCtrl THEN
           #FillingPhase.State.AutCtrl := FALSE;
           #FillingPhase.State.ManCtrl := TRUE;
           #FillingPhase.Cmd.ManCtrl := FALSE;
       END_IF;

       IF NOT #FillingPhase.State.AutCtrl AND NOT #FillingPhase.State.ManCtrl THEN
           #FillingPhase.State.ManCtrl := TRUE; // nebo dat Cmd.Manctrl do TRUE aby prosel IF nahore?
       END_IF;


    END_REGION

   REGION ManCtrl
       // processing manual actions - if command is processed, it is sets to FALSE even if can't be processed
       // Phase commands are start, stop, pause and resume 
       // Start - open filling valve 
       // Stop - close filling valve
       // Pause - close filling valve
       // Resume - open filling valve
       // real states of phase are writed into states in phase structure

       IF #FillingPhase.State.ManCtrl THEN
           IF #FillingPhase.Cmd.StartMan THEN
               #FillingPhase.State.Paused := FALSE;
               #FillingPhase.State.Idle := FALSE;
               #FillingPhase.State.Running := TRUE;

               #FillingValve.Cmd.OpenMan := TRUE;


               #FillingPhase.Cmd.ResetDone := TRUE;


           END_IF;

           IF #FillingPhase.State.Running THEN
               IF #FillingPhase.Cmd.PauseMan THEN
                   #FillingPhase.State.Running := FALSE;
                   #FillingPhase.State.Idle := FALSE;
                   #FillingPhase.State.Paused := TRUE;

                   #FillingValve.Cmd.CloseMan := TRUE;


                   #FillingPhase.Cmd.ResetDone := TRUE;

               END_IF;
           END_IF;

           IF #FillingPhase.State.Paused THEN
               IF #FillingPhase.Cmd.ResumeMan THEN
                   #FillingPhase.State.Paused := FALSE;
                   #FillingPhase.State.Idle := FALSE;
                   #FillingPhase.State.Running := TRUE;

                   #FillingValve.Cmd.OpenMan := TRUE;


                   #FillingPhase.Cmd.ResetDone := TRUE;

               END_IF;
           END_IF;


           IF #FillingPhase.State.Running OR #FillingPhase.State.Paused THEN
               IF #FillingPhase.Cmd.StopMan THEN
                   #FillingPhase.State.Running := FALSE;
                   #FillingPhase.State.Paused := FALSE;
                   #FillingPhase.State.Idle := TRUE;

                   #FillingValve.Cmd.CloseMan := TRUE;

                   #FillingPhase.Cmd.ResetDone := TRUE;


               END_IF;
           END_IF;



       END_IF;
       #FillingPhase.Cmd.StartMan := FALSE;
       #FillingPhase.Cmd.PauseMan := FALSE;
       #FillingPhase.Cmd.ResumeMan := FALSE;
       #FillingPhase.Cmd.StopMan := FALSE;



    END_REGION

   REGION AutCtrl
       // if request to run in automatic mode and phase can be run in automatic mode switch phase to running

       IF #FillingPhase.State.AutCtrl THEN
           IF #FillingPhase.Cmd.StartAut THEN
               #FillingPhase.State.Running := TRUE;
               #FillingPhase.State.Idle := FALSE;
               #FillingPhase.Cmd.StartAut := FALSE;
               #FillingValve.Cmd.AutCtrl := TRUE;
           END_IF;

           IF #FillingPhase.Cmd.StopAut THEN
               #FillingPhase.State.Running := FALSE;
               #FillingPhase.State.Idle := TRUE;
               #FillingPhase.Cmd.StopAut := FALSE;
           END_IF;

       END_IF;

    END_REGION

   REGION Done
       //every phase should have finish condition - filling phase - if water level is above requested level
       //after that done state should be setted to 1

       #FillingPhase.Param.FillLevel := 1.95;
       IF #FillingPhase.WaterLevel > #FillingPhase.Param.FillLevel THEN
           #FillingPhase.Cmd.StopAut := TRUE;
           #FillingPhase.Cmd.StopMan := TRUE;
           #FillingPhase.State.Done := TRUE;
       END_IF;

       // command reset done resets done state and than resets command

       IF #FillingPhase.Cmd.ResetDone THEN // AND DONE = TRUE? mozna zbytecne.
           #FillingPhase.State.Done := FALSE;
           #FillingPhase.Cmd.ResetDone := FALSE;
       END_IF;


       END_REGION

   REGION States 
       //Command valve in cases of states
       IF #FillingPhase.State.Running THEN
           #FillingValve.Cmd.Req2OpenAut := TRUE;
           #FillingValve.Cmd.Req2CloseAut := FALSE;
       ELSE
           #FillingValve.Cmd.Req2OpenAut := FALSE;
           #FillingValve.Cmd.Req2CloseAut := TRUE;
       END_IF;


       END_REGION


   // delault state of phase - if not any state sets state to idle
       IF NOT #FillingPhase.State.Idle AND NOT #FillingPhase.State.Paused AND NOT #FillingPhase.State.Running THEN
           #FillingPhase.State.Idle := TRUE;
   END_IF;

   // write binary states into int value for visualization

   IF #FillingPhase.State.Running THEN
       #FillingPhase.State.Stateint := #Running;
   ELSIF #FillingPhase.State.Paused THEN
       #FillingPhase.State.Stateint := #Pause;
   ELSIF #FillingPhase.State.Idle THEN
       #FillingPhase.State.Stateint := #Idle;
   ELSIF #FillingPhase.State.Done THEN
       #FillingPhase.State.Stateint := #Idle;
   END_IF;
END_FUNCTION_BLOCK

FUNCTION_BLOCK "DrainingFC"   // FB5, SCL
{ S7_Optimized_Access := 'TRUE' }
VERSION : 0.1
   VAR_IN_OUT
      DrainingPhase : "PhaseDraining";
      DrainingValve : "Valve";
   END_VAR
   VAR CONSTANT
      Idle : Int := 0;
      Running : Int := 1;
      Pause : Int := 2;
   END_VAR
BEGIN
   REGION Aut/Man
       // switching state of engine - automatic or manual control (default state is manual)
       IF #DrainingPhase.Cmd.AutCtrl THEN
           #DrainingPhase.State.ManCtrl := FALSE;
           #DrainingPhase.State.AutCtrl := TRUE;
           #DrainingPhase.Cmd.AutCtrl := FALSE;
       END_IF;

       IF #DrainingPhase.Cmd.ManCtrl THEN
           #DrainingPhase.State.AutCtrl := FALSE;
           #DrainingPhase.State.ManCtrl := TRUE;
           #DrainingPhase.Cmd.ManCtrl := FALSE;
       END_IF;

       IF NOT #DrainingPhase.State.AutCtrl AND NOT #DrainingPhase.State.ManCtrl THEN
           #DrainingPhase.State.ManCtrl := TRUE; // nebo dat Cmd.Manctrl do TRUE aby prosel IF nahore?
       END_IF;
   END_REGION

   REGION ManCtrl
       // processing manual actions - if command is processed, it is sets to FALSE even if can't be processed
       // Phase commands are start, stop, pause and resume 
       // Start - open draining valve 
       // Stop - close draining valve
       // Pause - close draining valve
       // Resume - open draining valve
       // real states of phase are writed into states in phase structure
       // 
       IF #DrainingPhase.State.ManCtrl THEN
           IF #DrainingPhase.Cmd.StartMan THEN
               #DrainingPhase.State.Paused := FALSE;
               #DrainingPhase.State.Idle := FALSE;
               #DrainingPhase.State.Running := TRUE;

               #DrainingValve.Cmd.OpenMan := TRUE; //?
               #DrainingValve.Cmd.OpenMan := FALSE;

               #DrainingPhase.Cmd.ResetDone := TRUE;
               #DrainingPhase.Cmd.ResetDone := FALSE;
           END_IF;

           IF #DrainingPhase.State.Running THEN
               IF #DrainingPhase.Cmd.PauseMan THEN
                   #DrainingPhase.State.Running := FALSE;
                   #DrainingPhase.State.Idle := FALSE;
                   #DrainingPhase.State.Paused := TRUE;

                   #DrainingValve.Cmd.CloseMan := TRUE;
                   #DrainingValve.Cmd.CloseMan := FALSE;

                   #DrainingPhase.Cmd.ResetDone := TRUE;
                   #DrainingPhase.Cmd.ResetDone := FALSE;
               END_IF;
           END_IF;

           IF #DrainingPhase.State.Paused THEN
               IF #DrainingPhase.Cmd.ResumeMan THEN
                   #DrainingPhase.State.Paused := FALSE;
                   #DrainingPhase.State.Idle := FALSE;
                   #DrainingPhase.State.Running := TRUE;

                   #DrainingValve.Cmd.OpenMan := TRUE;
                   #DrainingValve.Cmd.OpenMan := FALSE;

                   #DrainingPhase.Cmd.ResetDone := TRUE;
                   #DrainingPhase.Cmd.ResetDone := FALSE;
               END_IF;
           END_IF;


           IF #DrainingPhase.State.Running OR #DrainingPhase.State.Paused THEN
               IF #DrainingPhase.Cmd.StopMan THEN
                   #DrainingPhase.State.Running := FALSE;
                   #DrainingPhase.State.Paused := FALSE;
                   #DrainingPhase.State.Idle := TRUE;

                   #DrainingValve.Cmd.CloseMan := TRUE;
                   #DrainingValve.Cmd.CloseMan := FALSE;

                   #DrainingPhase.Cmd.ResetDone := TRUE;
                   #DrainingPhase.Cmd.ResetDone := FALSE;
               END_IF;
           END_IF;